REGION Network 17: Close Command
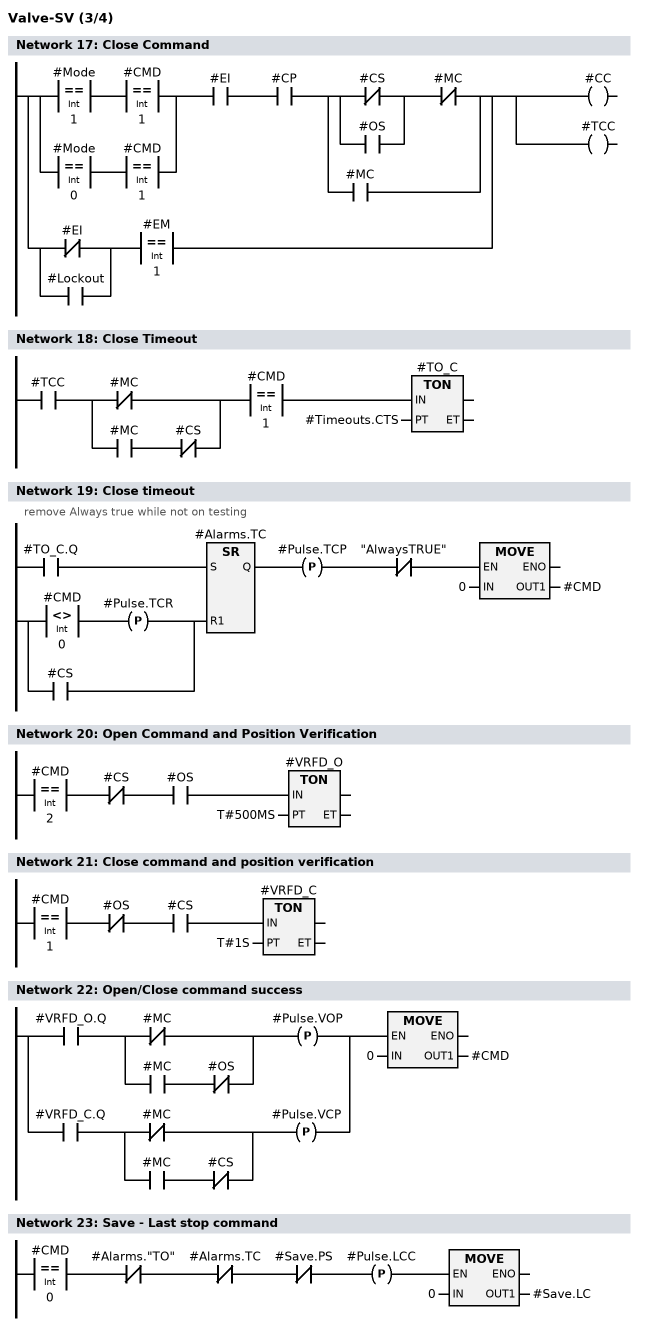
   RUNG wire#powerrail
      { S7_Templates := "SrcType := Int" } EQ_Contact(in1 := #Mode, in2 := 1)
      { S7_Templates := "SrcType := Int" } EQ_Contact(in1 := #CMD, in2 := 1)
      wire#w1
      Contact( #EI )
      Contact( #CP )
      wire#w2
      I_Contact( #CS )
      wire#w3
      I_Contact( #MC )
      wire#w4
      Coil( #CC )
   END_RUNG
   RUNG wire#powerrail
      { S7_Templates := "SrcType := Int" } EQ_Contact(in1 := #Mode, in2 := 0)
      { S7_Templates := "SrcType := Int" } EQ_Contact(in1 := #CMD, in2 := 1)
   END_RUNG wire#w1
   RUNG wire#w2
      Contact( #OS )
   END_RUNG wire#w3
   RUNG wire#w2
      Contact( #MC )
   END_RUNG wire#w4
   RUNG wire#powerrail
      I_Contact( #EI )
      wire#w5
      { S7_Templates := "SrcType := Int" } EQ_Contact(in1 := #EM, in2 := 1)
   END_RUNG wire#w4
   RUNG wire#powerrail
      Contact( #Lockout )
   END_RUNG wire#w5
   RUNG wire#w4
      Coil( #TCC )
   END_RUNG
   // the same network as SCL:
   #CC := ((((#Mode = 1) AND (#CMD = 1)) OR ((#Mode = 0) AND (#CMD = 1))) AND #EI AND #CP AND (((NOT #CS OR #OS) AND NOT #MC) OR #MC)) OR ((NOT #EI OR #Lockout) AND (#EM = 1));
   #TCC := #CC;
END_REGION

REGION Network 18: Close Timeout
   #TO_C(IN := #TCC AND (NOT #MC OR (#MC AND NOT #CS)) AND (#CMD = 1), PT := #Timeouts.CTS);   // TON
END_REGION

REGION Network 19: Close timeout
   // remove Always true while not on testing
   RUNG wire#powerrail
      Contact( #TO_C.Q )
      S_SR(operand := #Alarms.TC, r1 := wire#w1)
      P_Trig( #Pulse.TCP )
      I_Contact( "AlwaysTRUE" )
      { S7_GenerateENO := "TRUE" } Move(in := 0, out1 => #CMD)
   END_RUNG
   RUNG wire#powerrail
      { S7_Templates := "SrcType := Int" } NE_Contact(in1 := #CMD, in2 := 0)
      P_Trig( #Pulse.TCR )
   END_RUNG wire#w1
   RUNG wire#powerrail
      Contact( #CS )
   END_RUNG wire#w1
   // the same network as SCL:
   #_w1 := #CMD <> 0;
   #_w2 := #_w1 AND NOT #Pulse.TCR;   // rising edge
   #Pulse.TCR := #_w1;
   IF #TO_C.Q THEN
       #Alarms.TC := TRUE;   // SR flip-flop
   END_IF;
   IF #_w2 OR #CS THEN #Alarms.TC := FALSE; END_IF;
   #_w3 := #Alarms.TC AND NOT #Pulse.TCP;   // rising edge
   #Pulse.TCP := #Alarms.TC;
   IF #_w3 AND NOT "AlwaysTRUE" THEN #CMD := 0; END_IF;
END_REGION

REGION Network 20: Open Command and Position Verification
   #VRFD_O(IN := (#CMD = 2) AND NOT #CS AND #OS, PT := T#500MS);   // TON
END_REGION

REGION Network 21: Close command and position verification
   #VRFD_C(IN := (#CMD = 1) AND NOT #OS AND #CS, PT := T#1S);   // TON
END_REGION

REGION Network 22: Open/Close command success
   RUNG wire#powerrail
      Contact( #VRFD_O.Q )
      wire#w1
      I_Contact( #MC )
      wire#w2
      P_Trig( #Pulse.VOP )
      wire#w3
      { S7_GenerateENO := "TRUE" } Move(in := 0, out1 => #CMD)
   END_RUNG
   RUNG wire#w1
      Contact( #MC )
      I_Contact( #OS )
   END_RUNG wire#w2
   RUNG wire#powerrail
      Contact( #VRFD_C.Q )
      wire#w4
      I_Contact( #MC )
      wire#w5
      P_Trig( #Pulse.VCP )
   END_RUNG wire#w3
   RUNG wire#w4
      Contact( #MC )
      I_Contact( #CS )
   END_RUNG wire#w5
   // the same network as SCL:
   #_w1 := #VRFD_O.Q AND (NOT #MC OR (#MC AND NOT #OS));
   #_w2 := #_w1 AND NOT #Pulse.VOP;   // rising edge
   #Pulse.VOP := #_w1;
   #_w3 := #VRFD_C.Q AND (NOT #MC OR (#MC AND NOT #CS));
   #_w4 := #_w3 AND NOT #Pulse.VCP;   // rising edge
   #Pulse.VCP := #_w3;
   IF #_w2 OR #_w4 THEN #CMD := 0; END_IF;
END_REGION

REGION Network 23: Save - Last stop command
   RUNG wire#powerrail
      { S7_Templates := "SrcType := Int" } EQ_Contact(in1 := #CMD, in2 := 0)
      I_Contact( #Alarms."TO" )
      I_Contact( #Alarms.TC )
      I_Contact( #Save.PS )
      P_Trig( #Pulse.LCC )
      { S7_GenerateENO := "TRUE" } Move(in := 0, out1 => #Save.LC)
   END_RUNG
   // the same network as SCL:
   #_w1 := (#CMD = 0) AND NOT #Alarms."TO" AND NOT #Alarms.TC AND NOT #Save.PS;
   #_w2 := #_w1 AND NOT #Pulse.LCC;   // rising edge
   #Pulse.LCC := #_w1;
   IF #_w2 THEN #Save.LC := 0; END_IF;
END_REGION

REGION Network 24: Save - Last Stop Command
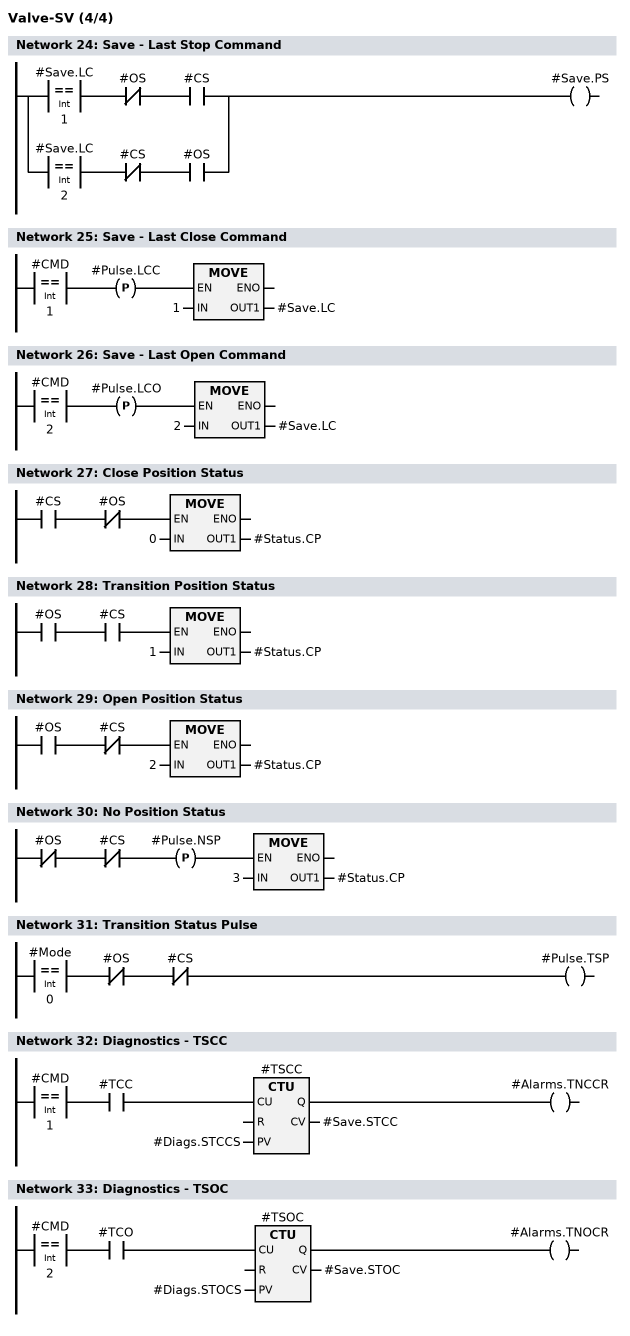
   RUNG wire#powerrail
      { S7_Templates := "SrcType := Int" } EQ_Contact(in1 := #Save.LC, in2 := 1)
      I_Contact( #OS )
      Contact( #CS )
      wire#w1
      Coil( #Save.PS )
   END_RUNG
   RUNG wire#powerrail
      { S7_Templates := "SrcType := Int" } EQ_Contact(in1 := #Save.LC, in2 := 2)
      I_Contact( #CS )
      Contact( #OS )
   END_RUNG wire#w1
   // the same network as SCL:
   #Save.PS := ((#Save.LC = 1) AND NOT #OS AND #CS) OR ((#Save.LC = 2) AND NOT #CS AND #OS);
END_REGION

REGION Network 25: Save - Last Close Command
   RUNG wire#powerrail
      { S7_Templates := "SrcType := Int" } EQ_Contact(in1 := #CMD, in2 := 1)
      P_Trig( #Pulse.LCC )
      { S7_GenerateENO := "TRUE" } Move(in := 1, out1 => #Save.LC)
   END_RUNG
   // the same network as SCL:
   #_w1 := #CMD = 1;
   #_w2 := #_w1 AND NOT #Pulse.LCC;   // rising edge
   #Pulse.LCC := #_w1;
   IF #_w2 THEN #Save.LC := 1; END_IF;
END_REGION

REGION Network 26: Save - Last Open Command
   RUNG wire#powerrail
      { S7_Templates := "SrcType := Int" } EQ_Contact(in1 := #CMD, in2 := 2)
      P_Trig( #Pulse.LCO )
      { S7_GenerateENO := "TRUE" } Move(in := 2, out1 => #Save.LC)
   END_RUNG
   // the same network as SCL:
   #_w1 := #CMD = 2;
   #_w2 := #_w1 AND NOT #Pulse.LCO;   // rising edge
   #Pulse.LCO := #_w1;
   IF #_w2 THEN #Save.LC := 2; END_IF;
END_REGION

REGION Network 27: Close Position Status
   RUNG wire#powerrail
      Contact( #CS )
      I_Contact( #OS )
      { S7_GenerateENO := "TRUE" } Move(in := 0, out1 => #Status.CP)
   END_RUNG
   // the same network as SCL:
   IF #CS AND NOT #OS THEN #Status.CP := 0; END_IF;
END_REGION

REGION Network 28: Transition Position Status
   RUNG wire#powerrail
      Contact( #OS )
      Contact( #CS )
      { S7_GenerateENO := "TRUE" } Move(in := 1, out1 => #Status.CP)
   END_RUNG
   // the same network as SCL:
   IF #OS AND #CS THEN #Status.CP := 1; END_IF;
END_REGION

REGION Network 29: Open Position Status
   RUNG wire#powerrail
      Contact( #OS )
      I_Contact( #CS )
      { S7_GenerateENO := "TRUE" } Move(in := 2, out1 => #Status.CP)
   END_RUNG
   // the same network as SCL:
   IF #OS AND NOT #CS THEN #Status.CP := 2; END_IF;
END_REGION

REGION Network 30: No Position Status
   RUNG wire#powerrail
      I_Contact( #OS )
      I_Contact( #CS )
      P_Trig( #Pulse.NSP )
      { S7_GenerateENO := "TRUE" } Move(in := 3, out1 => #Status.CP)
   END_RUNG
   // the same network as SCL:
   #_w1 := NOT #OS AND NOT #CS;
   #_w2 := #_w1 AND NOT #Pulse.NSP;   // rising edge
   #Pulse.NSP := #_w1;
   IF #_w2 THEN #Status.CP := 3; END_IF;
END_REGION

REGION Network 31: Transition Status Pulse
   RUNG wire#powerrail
      { S7_Templates := "SrcType := Int" } EQ_Contact(in1 := #Mode, in2 := 0)
      I_Contact( #OS )
      I_Contact( #CS )
      Coil( #Pulse.TSP )
   END_RUNG
   // the same network as SCL:
   #Pulse.TSP := (#Mode = 0) AND NOT #OS AND NOT #CS;
END_REGION

REGION Network 32: Diagnostics - TSCC
   #TSCC(CU := (#CMD = 1) AND #TCC, PV := #Diags.STCCS, CV => #Save.STCC);   // CTU
   #Alarms.TNCCR := #TSCC.Q;
END_REGION

REGION Network 33: Diagnostics - TSOC
   #TSOC(CU := (#CMD = 2) AND #TCO, PV := #Diags.STOCS, CV => #Save.STOC);   // CTU
   #Alarms.TNOCR := #TSOC.Q;
END_REGION
END_FUNCTION_BLOCK

FUNCTION_BLOCK "Valve-CV"   // FB801, LAD
TITLE = Valve-CV
{ S7_Optimized_Access := 'TRUE' }
VERSION : 0.1
// V1.0    GE    04/04/2022     Modified Unscale block and made sure CMD outputs right number.
   VAR_INPUT
      POS_CMD_Word : Word;   // Command in Word
      POS_FB : Int;   // Valve Position Raw Value
      AnalogFeedbackExists : Bool;   // Feedback Mode FALSE=FDBK Off // TRUE=FDBCK On
   END_VAR
   VAR_OUTPUT
      CMD : Int;   // Commanded Position in INT format
      CMD_R : Real;
   END_VAR
   VAR
      HMI : Struct
         Controls : Struct   // Controls
            SP : Real;   // Operator Command
            Lockout : Bool;
         END_STRUCT;
         Status : Struct   // Status
            POS : Real;   // Valve Position
            LST_POS : Real;   // Valve Position after a successful transition
            CMD_SP : Real;   // Commanded Position
            WR : Bool;   // Within Range
            UR_DB : Real;   // Upper range deadband
            LR_DB : Real;   // Lower range Deadband
            Mode_A : Bool;
            Mode_B : Bool;
         END_STRUCT;
         Alarms : Struct
            FCMD : Bool;   // SP vs PV mismatch timeout
            SP : Real;   // Setpoint Alarm (Unused)
            Error : Word;   // Unscaling Error
            IL : Bool := TRUE ;   // INTERLOCK (TRUE= GOOD FALSE = BAD)
         END_STRUCT;
         Config : Struct
            Mode : Int;   // 0 = PLC, 1 = HMI
            FDBK_MD : Int;   // Feedback Mode 0=FDBK Off // 1=FDBCK On
            WR_DB_TON : Time := T#1S;   // PV within range of SP
            WR_DB_TOF : Time := T#1S;   // PV within range of SP
            CMD_TO_TON_PT : Time := T#10S;   // Command to Open TON Preset Time
            CMD_TO_TOF_PT : Time := T#1S;   // Command to Open TOF Preset Time
            UR_DB_SP : Real := 1.0;   // Upper Range Deadband Setpoint
            LR_DB_SP : Real := 1.0;   // Lower Range Deadband Setpoint
            Min : Real;   // Minimum Output
            Max : Real := 100.0;   // Max Output
            failOpen : Bool;   // Enable Bipolar Values in Control Value
         END_STRUCT;
      END_STRUCT;
      OS : Struct
         SaveLastSP : Bool;   // Save Last Valid Setpoint
      END_STRUCT;
      WR_DB_TON : TON_TIME;   // Within Range Debounce TON
      WR_DB_TOF : TOF_TIME;   // Withing Range Debounce TOF
      CMD_TO_TON : TON_TIME;   // Command Timeout Debounce
      CMD_TO_TOF : TOF_TIME;   // Command Timeout Debounce
      "Lockout Trig" : Bool;
   END_VAR
   VAR_TEMP
      Scale : Struct
         RAI : Real;   // CV Position in REAL data type format
         EMax : Real;   // Engineering Max
         EMin : Real;   // Engineering Min
         RMax : Real;   // Raw Max
         RMin : Real;   // Raw Max
         OFST : Real;   // Offset
         RRAnge : Real;   // Raw Range
         ERange : Real;   // Engineering Range
      END_STRUCT;
      RDI : DInt;
      M1 : Real;
      M2 : Real;
      M3 : Real;
      CMD_SP : Real;
      WR : Bool;
      WR_DB : Bool;
      FCMD : Bool;   // SP vs PV mismatch timeout
      bypass : Bool;
      NRAIR : Real;
   END_VAR
   VAR_TEMP   // added for the SCL form of the ladder/FBD networks
      _w1 : Bool;
   END_VAR
BEGIN

REGION Network 1: Feedback MODE
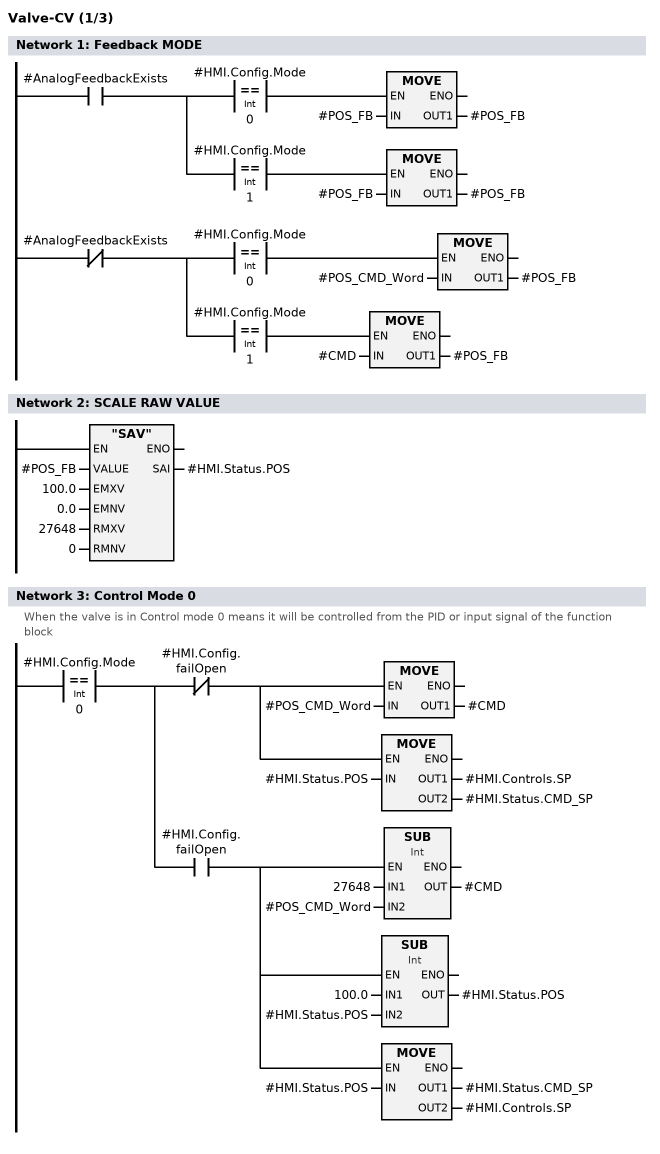
   RUNG wire#powerrail
      Contact( #AnalogFeedbackExists )
      wire#w1
      { S7_Templates := "SrcType := Int" } EQ_Contact(in1 := #HMI.Config.Mode, in2 := 0)
      Move(in := #POS_FB, out1 => #POS_FB)
   END_RUNG
   RUNG wire#w1
      { S7_Templates := "SrcType := Int" } EQ_Contact(in1 := #HMI.Config.Mode, in2 := 1)
      Move(in := #POS_FB, out1 => #POS_FB)
   END_RUNG
   RUNG wire#powerrail
      I_Contact( #AnalogFeedbackExists )
      wire#w2
      { S7_Templates := "SrcType := Int" } EQ_Contact(in1 := #HMI.Config.Mode, in2 := 0)
      Move(in := #POS_CMD_Word, out1 => #POS_FB)
   END_RUNG
   RUNG wire#w2
      { S7_Templates := "SrcType := Int" } EQ_Contact(in1 := #HMI.Config.Mode, in2 := 1)
      Move(in := #CMD, out1 => #POS_FB)
   END_RUNG
   // the same network as SCL:
   IF #AnalogFeedbackExists AND (#HMI.Config.Mode = 0) THEN #POS_FB := #POS_FB; END_IF;
   IF #AnalogFeedbackExists AND (#HMI.Config.Mode = 1) THEN #POS_FB := #POS_FB; END_IF;
   #_w1 := NOT #AnalogFeedbackExists;
   IF #_w1 AND (#HMI.Config.Mode = 0) THEN #POS_FB := #POS_CMD_Word; END_IF;
   IF #_w1 AND (#HMI.Config.Mode = 1) THEN #POS_FB := #CMD; END_IF;
END_REGION

REGION Network 2: SCALE RAW VALUE
   RUNG wire#powerrail
      "SAV"(VALUE := #POS_FB, EMXV := 100.0, EMNV := 0.0, RMXV := 27648, RMNV := 0, SAI => #HMI.Status.POS)
   END_RUNG
   // the same network as SCL:
   "SAV"(VALUE := #POS_FB, EMXV := 100.0, EMNV := 0.0, RMXV := 27648, RMNV := 0, SAI => #HMI.Status.POS);
END_REGION

REGION Network 3: Control Mode 0
   // When the valve is in Control mode 0 means it will be controlled from the PID or input signal of the function block
   RUNG wire#powerrail
      { S7_Templates := "SrcType := Int" } EQ_Contact(in1 := #HMI.Config.Mode, in2 := 0)
      wire#w1
      I_Contact( #HMI.Config.failOpen )
      wire#w2
      { S7_GenerateENO := "TRUE" } Move(in := #POS_CMD_Word, out1 => #CMD)
   END_RUNG
   RUNG wire#w2
      Move(in := #HMI.Status.POS, out1 => #HMI.Controls.SP, out2 => #HMI.Status.CMD_SP)
   END_RUNG
   RUNG wire#w1
      Contact( #HMI.Config.failOpen )
      wire#w3
      { S7_Templates := "SrcType := Int" } Sub(in1 := 27648, in2 := #POS_CMD_Word, out => #CMD)
   END_RUNG
   RUNG wire#w3
      { S7_Templates := "SrcType := Int" } Sub(in1 := 100.0, in2 := #HMI.Status.POS, out => #HMI.Status.POS)
   END_RUNG
   RUNG wire#w3
      Move(in := #HMI.Status.POS, out1 => #HMI.Status.CMD_SP, out2 => #HMI.Controls.SP)
   END_RUNG
   // the same network as SCL:
   #_w1 := #HMI.Config.Mode = 0;
   IF #_w1 AND NOT #HMI.Config.failOpen THEN
       #CMD := #POS_CMD_Word;
       #HMI.Controls.SP := #HMI.Status.POS;
       #HMI.Status.CMD_SP := #HMI.Status.POS;
   END_IF;
   IF #_w1 AND #HMI.Config.failOpen THEN
       #CMD := 27648 - #POS_CMD_Word;
       #HMI.Status.POS := 100.0 - #HMI.Status.POS;
       #HMI.Status.CMD_SP := #HMI.Status.POS;
       #HMI.Controls.SP := #HMI.Status.POS;
   END_IF;
END_REGION

REGION Network 4: Control Mode 1
   // Control Mode 1 will control from HMI (force valve to go to a certain position)
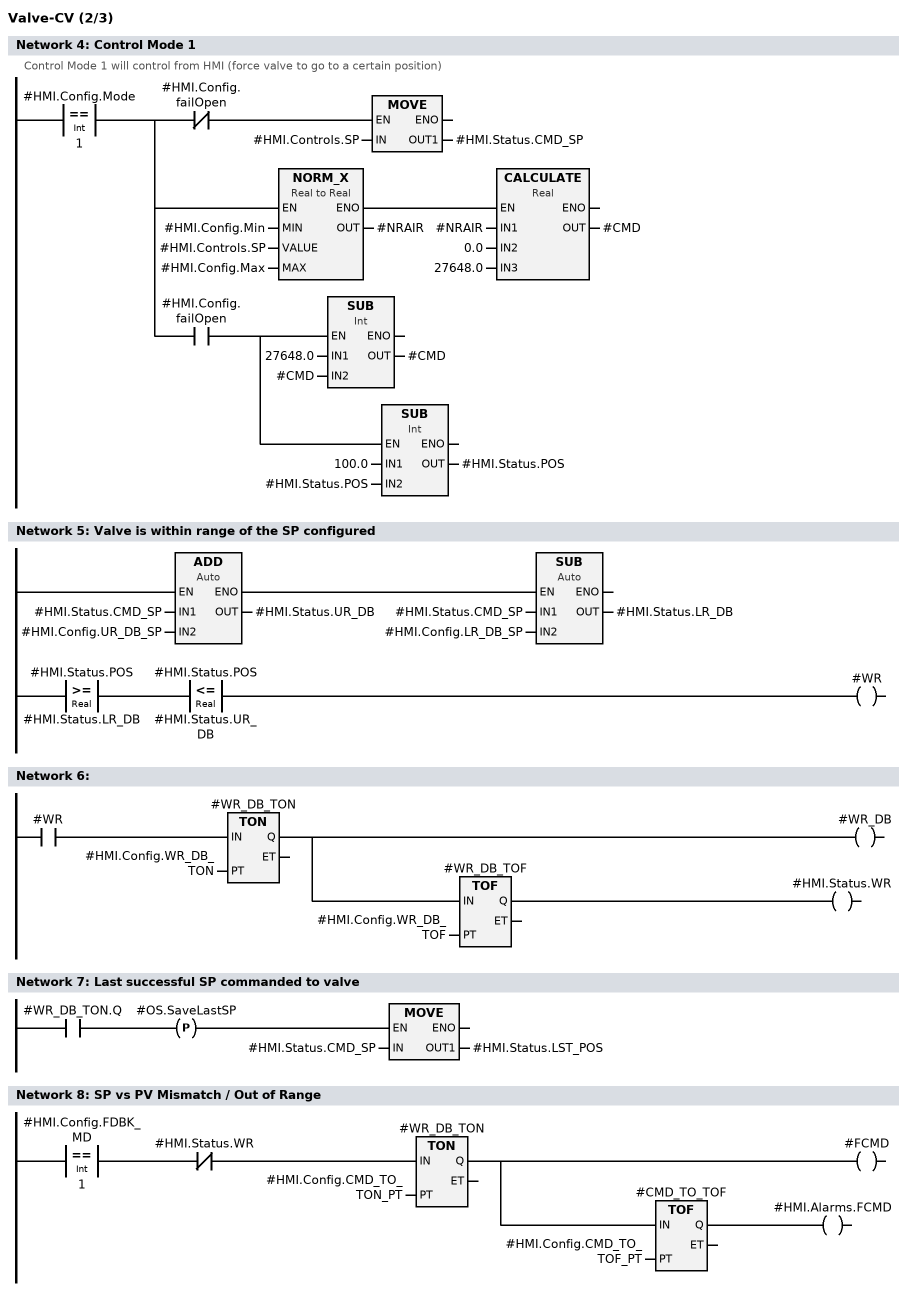
   RUNG wire#powerrail
      { S7_Templates := "SrcType := Int" } EQ_Contact(in1 := #HMI.Config.Mode, in2 := 1)
      wire#w1
      I_Contact( #HMI.Config.failOpen )
      { S7_GenerateENO := "TRUE" } Move(in := #HMI.Controls.SP, out1 => #HMI.Status.CMD_SP)
   END_RUNG
   RUNG wire#w1
      { S7_Templates := "[SrcType := Real, DestType := Real]" } Normalize(min := #HMI.Config.Min, value := #HMI.Controls.SP, max := #HMI.Config.Max, out => #NRAIR)
      { S7_Templates := "SrcType := Real"; S7_Expression := "(IN1 * (IN3 - IN2)) + IN2" } Calculate(in1 := #NRAIR, in2 := 0.0, in3 := 27648.0, out => #CMD)
   END_RUNG
   RUNG wire#w1
      Contact( #HMI.Config.failOpen )
      wire#w2
      { S7_Templates := "SrcType := Int" } Sub(in1 := 27648.0, in2 := #CMD, out => #CMD)
   END_RUNG
   RUNG wire#w2
      { S7_Templates := "SrcType := Int" } Sub(in1 := 100.0, in2 := #HMI.Status.POS, out => #HMI.Status.POS)
   END_RUNG
   // the same network as SCL:
   #_w1 := #HMI.Config.Mode = 1;
   IF #_w1 AND NOT #HMI.Config.failOpen THEN #HMI.Status.CMD_SP := #HMI.Controls.SP; END_IF;
   IF #_w1 THEN
       #NRAIR := NORM_X(MIN := #HMI.Config.Min, VALUE := #HMI.Controls.SP, MAX := #HMI.Config.Max);
       #CMD := (#NRAIR * (27648.0 - 0.0)) + 0.0;
   END_IF;
   IF #_w1 AND #HMI.Config.failOpen THEN
       #CMD := 27648.0 - #CMD;
       #HMI.Status.POS := 100.0 - #HMI.Status.POS;
   END_IF;
END_REGION

REGION Network 5: Valve is within range of the SP configured
   RUNG wire#powerrail
      Add(in1 := #HMI.Status.CMD_SP, in2 := #HMI.Config.UR_DB_SP, out => #HMI.Status.UR_DB)
      Sub(in1 := #HMI.Status.CMD_SP, in2 := #HMI.Config.LR_DB_SP, out => #HMI.Status.LR_DB)
   END_RUNG
   RUNG wire#powerrail
      { S7_Templates := "SrcType := Real" } GE_Contact(in1 := #HMI.Status.POS, in2 := #HMI.Status.LR_DB)
      { S7_Templates := "SrcType := Real" } LE_Contact(in1 := #HMI.Status.POS, in2 := #HMI.Status.UR_DB)
      Coil( #WR )
   END_RUNG
   // the same network as SCL:
   #HMI.Status.UR_DB := #HMI.Status.CMD_SP + #HMI.Config.UR_DB_SP;
   #HMI.Status.LR_DB := #HMI.Status.CMD_SP - #HMI.Config.LR_DB_SP;
   #WR := (#HMI.Status.POS >= #HMI.Status.LR_DB) AND (#HMI.Status.POS <= #HMI.Status.UR_DB);
END_REGION

REGION Network 6
   #WR_DB_TON(IN := #WR, PT := #HMI.Config.WR_DB_TON);   // TON
   #WR_DB := #WR_DB_TON.Q;
   #WR_DB_TOF(IN := #WR_DB_TON.Q, PT := #HMI.Config.WR_DB_TOF);   // TOF
   #HMI.Status.WR := #WR_DB_TOF.Q;
END_REGION

REGION Network 7: Last successful SP commanded to valve
   RUNG wire#powerrail
      Contact( #WR_DB_TON.Q )
      P_Trig( #OS.SaveLastSP )
      { S7_GenerateENO := "TRUE" } Move(in := #HMI.Status.CMD_SP, out1 => #HMI.Status.LST_POS)
   END_RUNG
   // the same network as SCL:
   #_w1 := #WR_DB_TON.Q AND NOT #OS.SaveLastSP;   // rising edge
   #OS.SaveLastSP := #WR_DB_TON.Q;
   IF #_w1 THEN #HMI.Status.LST_POS := #HMI.Status.CMD_SP; END_IF;
END_REGION

REGION Network 8: SP vs PV Mismatch / Out of Range
   #WR_DB_TON(IN := (#HMI.Config.FDBK_MD = 1) AND NOT #HMI.Status.WR, PT := #HMI.Config.CMD_TO_TON_PT);   // TON
   #FCMD := #WR_DB_TON.Q;
   #CMD_TO_TOF(IN := #WR_DB_TON.Q, PT := #HMI.Config.CMD_TO_TOF_PT);   // TOF
   #HMI.Alarms.FCMD := #CMD_TO_TOF.Q;
END_REGION

REGION Network 9: Lockout Sequence
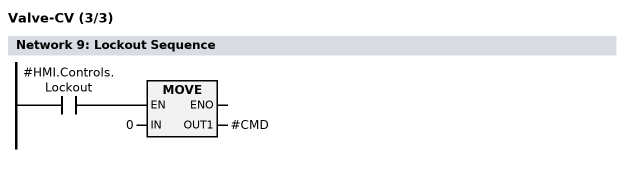
   RUNG wire#powerrail
      Contact( #HMI.Controls.Lockout )
      { S7_GenerateENO := "TRUE" } Move(in := 0, out1 => #CMD)
   END_RUNG
   // the same network as SCL:
   IF #HMI.Controls.Lockout THEN #CMD := 0; END_IF;
END_REGION
END_FUNCTION_BLOCK

// folder: Analogs inputs

FUNCTION "Analog Trasmitter" : Void   // FC5, LAD
TITLE = Analog Trasmitter Fuction Code
{ S7_Optimized_Access := 'TRUE' }
VERSION : 0.1
// Updated Date:
// Note:
BEGIN
END_FUNCTION

// folder: Analogs inputs/Trasmitters/Analyzer Trasmitters

FUNCTION "Analyzer Trasmitters" : Void   // FC16, LAD
TITLE = Analyzer Trasmitters
{ S7_Optimized_Access := 'TRUE' }
VERSION : 0.1
// Updated Date:
// Note:
BEGIN

REGION Network 1: AT-3011 : C-301 Nitrates Analyzer #1
   // Erick
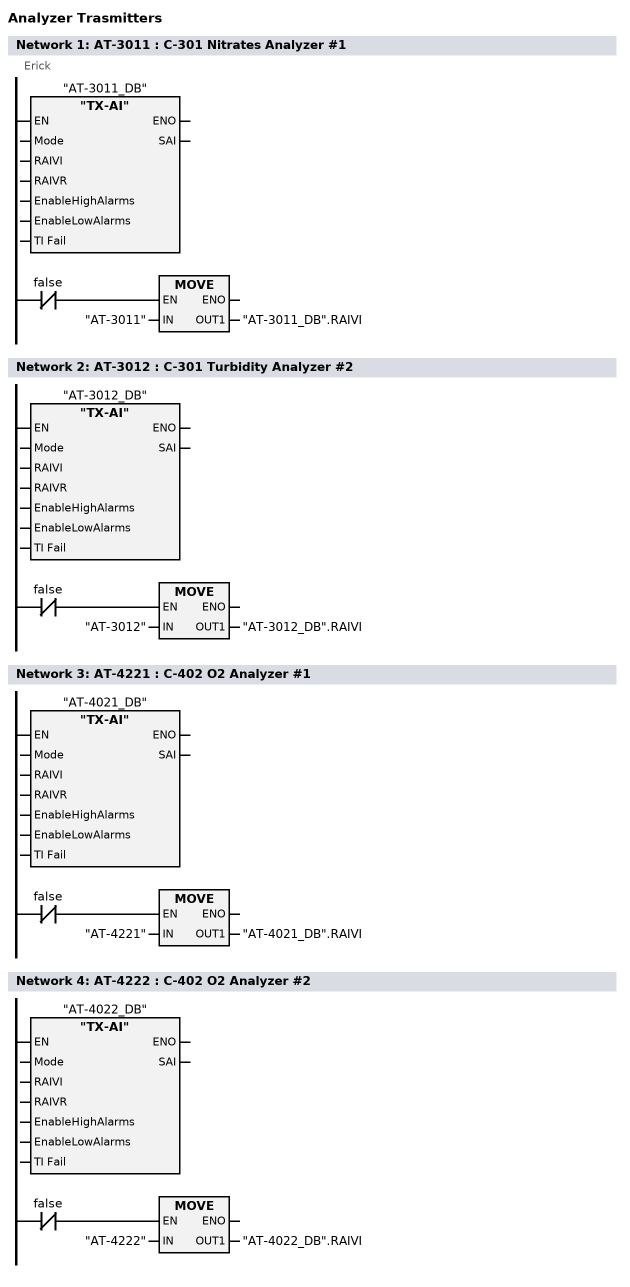
   RUNG wire#powerrail
      "AT-3011_DB"(Mode :=, RAIVI :=, RAIVR :=, EnableHighAlarms :=, EnableLowAlarms :=, "TI Fail" :=, SAI =>)
   END_RUNG
   RUNG wire#powerrail
      I_Contact( false )
      { S7_GenerateENO := "TRUE" } Move(in := "AT-3011", out1 => "AT-3011_DB".RAIVI)
   END_RUNG
   // the same network as SCL:
   "AT-3011_DB"();   // "TX-AI"
   IF NOT false THEN "AT-3011_DB".RAIVI := "AT-3011"; END_IF;
END_REGION

REGION Network 2: AT-3012 : C-301 Turbidity Analyzer #2
   RUNG wire#powerrail
      "AT-3012_DB"(Mode :=, RAIVI :=, RAIVR :=, EnableHighAlarms :=, EnableLowAlarms :=, "TI Fail" :=, SAI =>)
   END_RUNG
   RUNG wire#powerrail
      I_Contact( false )
      { S7_GenerateENO := "TRUE" } Move(in := "AT-3012", out1 => "AT-3012_DB".RAIVI)
   END_RUNG
   // the same network as SCL:
   "AT-3012_DB"();   // "TX-AI"
   IF NOT false THEN "AT-3012_DB".RAIVI := "AT-3012"; END_IF;
END_REGION

REGION Network 3: AT-4221 : C-402 O2 Analyzer #1
   RUNG wire#powerrail
      "AT-4021_DB"(Mode :=, RAIVI :=, RAIVR :=, EnableHighAlarms :=, EnableLowAlarms :=, "TI Fail" :=, SAI =>)
   END_RUNG
   RUNG wire#powerrail
      I_Contact( false )
      { S7_GenerateENO := "TRUE" } Move(in := "AT-4221", out1 => "AT-4021_DB".RAIVI)
   END_RUNG
   // the same network as SCL:
   "AT-4021_DB"();   // "TX-AI"
   IF NOT false THEN "AT-4021_DB".RAIVI := "AT-4221"; END_IF;
END_REGION

REGION Network 4: AT-4222 : C-402 O2 Analyzer #2
   RUNG wire#powerrail
      "AT-4022_DB"(Mode :=, RAIVI :=, RAIVR :=, EnableHighAlarms :=, EnableLowAlarms :=, "TI Fail" :=, SAI =>)
   END_RUNG
   RUNG wire#powerrail
      I_Contact( false )
      { S7_GenerateENO := "TRUE" } Move(in := "AT-4222", out1 => "AT-4022_DB".RAIVI)
   END_RUNG
   // the same network as SCL:
   "AT-4022_DB"();   // "TX-AI"
   IF NOT false THEN "AT-4022_DB".RAIVI := "AT-4222"; END_IF;
END_REGION
END_FUNCTION

// folder: Analogs inputs/Trasmitters/Flow Trasmitters

FUNCTION "FlowTrasmitters" : Void   // FC8, LAD
TITLE = Flow Trasmitter Fuction Code
{ S7_Optimized_Access := 'TRUE' }
VERSION : 0.1
// Updated Date:
// Note:
BEGIN

REGION Network 1: FT-1011: T-101 Recirc Flow
   // "FT-1011"
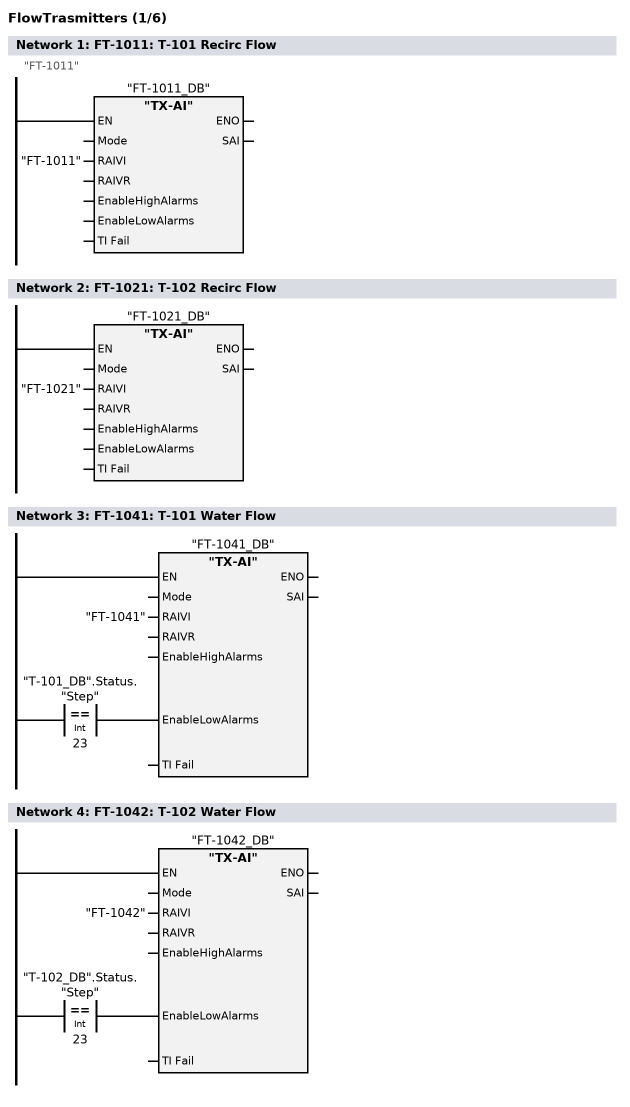
   RUNG wire#powerrail
      "FT-1011_DB"(Mode :=, RAIVI := "FT-1011", RAIVR :=, EnableHighAlarms :=, EnableLowAlarms :=, "TI Fail" :=, SAI =>)
   END_RUNG
   // the same network as SCL:
   "FT-1011_DB"(RAIVI := "FT-1011");   // "TX-AI"
END_REGION

REGION Network 2: FT-1021: T-102 Recirc Flow
   RUNG wire#powerrail
      "FT-1021_DB"(Mode :=, RAIVI := "FT-1021", RAIVR :=, EnableHighAlarms :=, EnableLowAlarms :=, "TI Fail" :=, SAI =>)
   END_RUNG
   // the same network as SCL:
   "FT-1021_DB"(RAIVI := "FT-1021");   // "TX-AI"
END_REGION

REGION Network 3: FT-1041: T-101 Water Flow
   RUNG wire#powerrail
      "FT-1041_DB"(EnableLowAlarms := wire#w1, Mode :=, RAIVI := "FT-1041", RAIVR :=, EnableHighAlarms :=, "TI Fail" :=, SAI =>)
   END_RUNG
   RUNG wire#powerrail
      { S7_Templates := "SrcType := Int" } EQ_Contact(in1 := "T-101_DB".Status."Step", in2 := 23)
   END_RUNG wire#w1
   // the same network as SCL:
   "FT-1041_DB"(RAIVI := "FT-1041", EnableLowAlarms := "T-101_DB".Status."Step" = 23);   // "TX-AI"
END_REGION

REGION Network 4: FT-1042: T-102 Water Flow
   RUNG wire#powerrail
      "FT-1042_DB"(EnableLowAlarms := wire#w1, Mode :=, RAIVI := "FT-1042", RAIVR :=, EnableHighAlarms :=, "TI Fail" :=, SAI =>)
   END_RUNG
   RUNG wire#powerrail
      { S7_Templates := "SrcType := Int" } EQ_Contact(in1 := "T-102_DB".Status."Step", in2 := 23)
   END_RUNG wire#w1
   // the same network as SCL:
   "FT-1042_DB"(RAIVI := "FT-1042", EnableLowAlarms := "T-102_DB".Status."Step" = 23);   // "TX-AI"
END_REGION

REGION Network 5: FT-1043:R-201 Water Flow
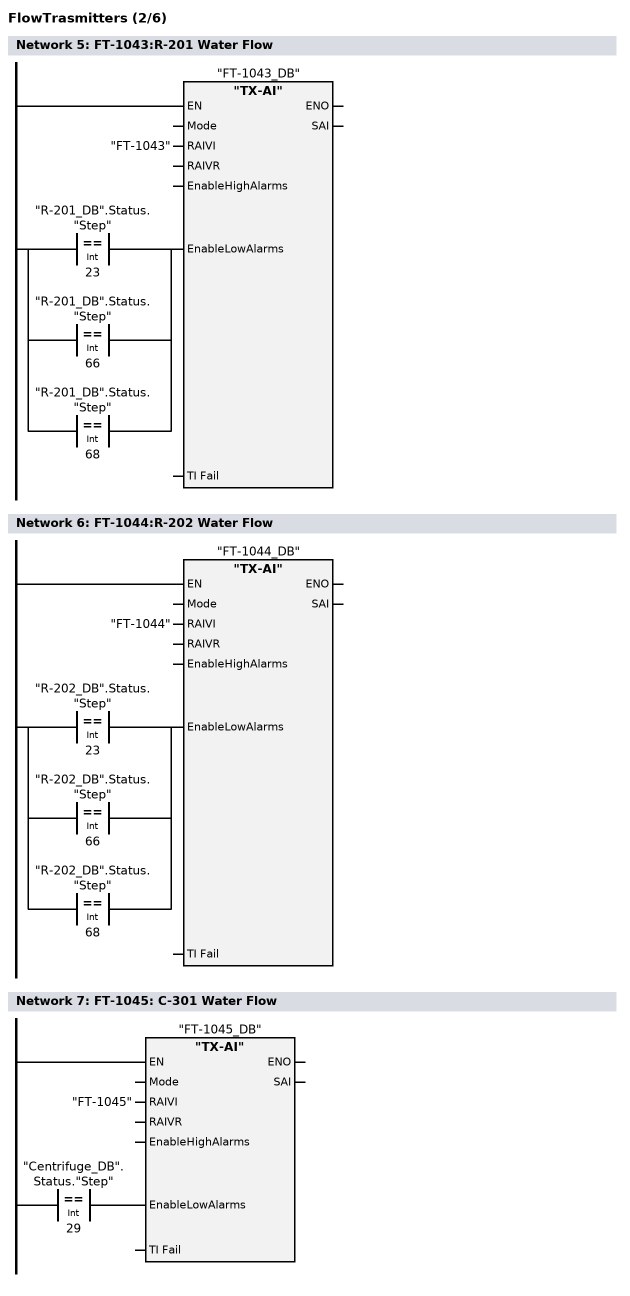
   RUNG wire#powerrail
      "FT-1043_DB"(EnableLowAlarms := wire#w1, Mode :=, RAIVI := "FT-1043", RAIVR :=, EnableHighAlarms :=, "TI Fail" :=, SAI =>)
   END_RUNG
   RUNG wire#powerrail
      { S7_Templates := "SrcType := Int" } EQ_Contact(in1 := "R-201_DB".Status."Step", in2 := 23)
   END_RUNG wire#w1
   RUNG wire#powerrail
      { S7_Templates := "SrcType := Int" } EQ_Contact(in1 := "R-201_DB".Status."Step", in2 := 66)
   END_RUNG wire#w1
   RUNG wire#powerrail
      { S7_Templates := "SrcType := Int" } EQ_Contact(in1 := "R-201_DB".Status."Step", in2 := 68)
   END_RUNG wire#w1
   // the same network as SCL:
   "FT-1043_DB"(RAIVI := "FT-1043",   // "TX-AI"
                EnableLowAlarms := ("R-201_DB".Status."Step" = 23) OR ("R-201_DB".Status."Step" = 66) OR ("R-201_DB".Status."Step" = 68));
END_REGION

REGION Network 6: FT-1044:R-202 Water Flow
   RUNG wire#powerrail
      "FT-1044_DB"(EnableLowAlarms := wire#w1, Mode :=, RAIVI := "FT-1044", RAIVR :=, EnableHighAlarms :=, "TI Fail" :=, SAI =>)
   END_RUNG
   RUNG wire#powerrail
      { S7_Templates := "SrcType := Int" } EQ_Contact(in1 := "R-202_DB".Status."Step", in2 := 23)
   END_RUNG wire#w1
   RUNG wire#powerrail
      { S7_Templates := "SrcType := Int" } EQ_Contact(in1 := "R-202_DB".Status."Step", in2 := 66)
   END_RUNG wire#w1
   RUNG wire#powerrail
      { S7_Templates := "SrcType := Int" } EQ_Contact(in1 := "R-202_DB".Status."Step", in2 := 68)
   END_RUNG wire#w1
   // the same network as SCL:
   "FT-1044_DB"(RAIVI := "FT-1044",   // "TX-AI"
                EnableLowAlarms := ("R-202_DB".Status."Step" = 23) OR ("R-202_DB".Status."Step" = 66) OR ("R-202_DB".Status."Step" = 68));
END_REGION

REGION Network 7: FT-1045: C-301 Water Flow
   RUNG wire#powerrail
      "FT-1045_DB"(EnableLowAlarms := wire#w1, Mode :=, RAIVI := "FT-1045", RAIVR :=, EnableHighAlarms :=, "TI Fail" :=, SAI =>)
   END_RUNG
   RUNG wire#powerrail
      { S7_Templates := "SrcType := Int" } EQ_Contact(in1 := "Centrifuge_DB".Status."Step", in2 := 29)
   END_RUNG wire#w1
   // the same network as SCL:
   "FT-1045_DB"(RAIVI := "FT-1045", EnableLowAlarms := "Centrifuge_DB".Status."Step" = 29);   // "TX-AI"
END_REGION

REGION Network 8: FT-2011:T-101 to R-201 Flow
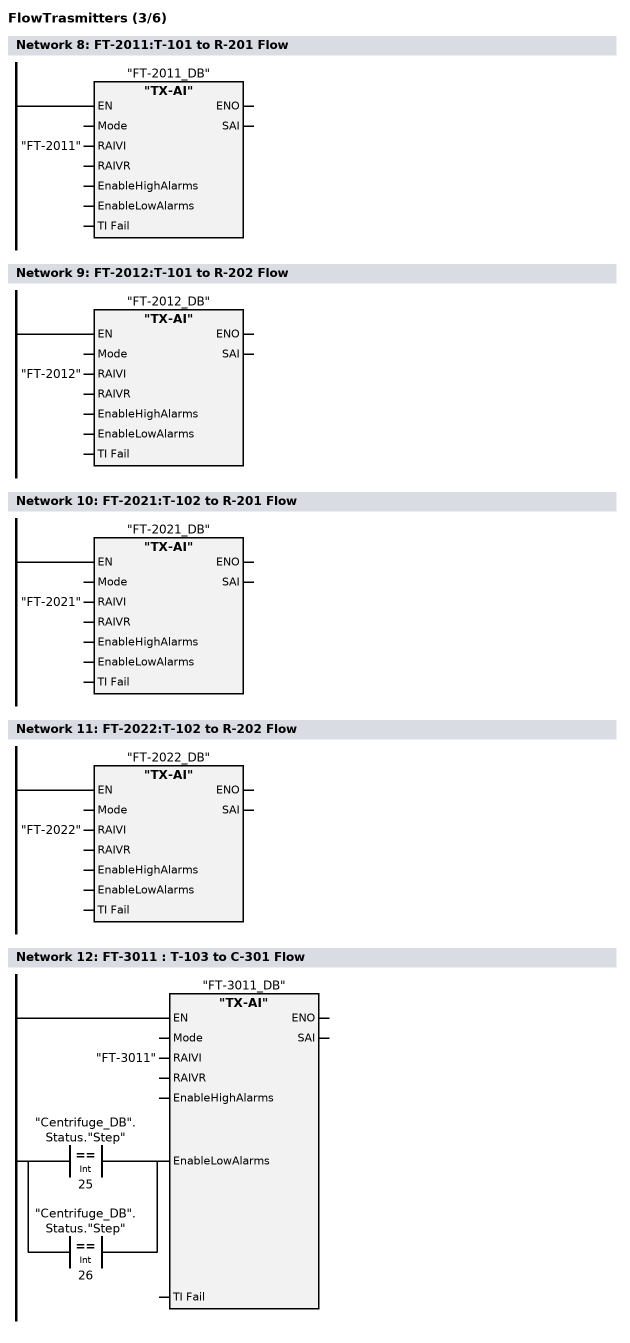
   RUNG wire#powerrail
      "FT-2011_DB"(Mode :=, RAIVI := "FT-2011", RAIVR :=, EnableHighAlarms :=, EnableLowAlarms :=, "TI Fail" :=, SAI =>)
   END_RUNG
   // the same network as SCL:
   "FT-2011_DB"(RAIVI := "FT-2011");   // "TX-AI"
END_REGION

REGION Network 9: FT-2012:T-101 to R-202 Flow
   RUNG wire#powerrail
      "FT-2012_DB"(Mode :=, RAIVI := "FT-2012", RAIVR :=, EnableHighAlarms :=, EnableLowAlarms :=, "TI Fail" :=, SAI =>)
   END_RUNG
   // the same network as SCL:
   "FT-2012_DB"(RAIVI := "FT-2012");   // "TX-AI"
END_REGION

REGION Network 10: FT-2021:T-102 to R-201 Flow
   RUNG wire#powerrail
      "FT-2021_DB"(Mode :=, RAIVI := "FT-2021", RAIVR :=, EnableHighAlarms :=, EnableLowAlarms :=, "TI Fail" :=, SAI =>)
   END_RUNG
   // the same network as SCL:
   "FT-2021_DB"(RAIVI := "FT-2021");   // "TX-AI"
END_REGION

REGION Network 11: FT-2022:T-102 to R-202 Flow
   RUNG wire#powerrail
      "FT-2022_DB"(Mode :=, RAIVI := "FT-2022", RAIVR :=, EnableHighAlarms :=, EnableLowAlarms :=, "TI Fail" :=, SAI =>)
   END_RUNG
   // the same network as SCL:
   "FT-2022_DB"(RAIVI := "FT-2022");   // "TX-AI"
END_REGION

REGION Network 12: FT-3011 : T-103 to C-301 Flow
   RUNG wire#powerrail
      "FT-3011_DB"(EnableLowAlarms := wire#w1, Mode :=, RAIVI := "FT-3011", RAIVR :=, EnableHighAlarms :=, "TI Fail" :=, SAI =>)
   END_RUNG
   RUNG wire#powerrail
      { S7_Templates := "SrcType := Int" } EQ_Contact(in1 := "Centrifuge_DB".Status."Step", in2 := 25)
   END_RUNG wire#w1
   RUNG wire#powerrail
      { S7_Templates := "SrcType := Int" } EQ_Contact(in1 := "Centrifuge_DB".Status."Step", in2 := 26)
   END_RUNG wire#w1
   // the same network as SCL:
   "FT-3011_DB"(RAIVI := "FT-3011",   // "TX-AI"
                EnableLowAlarms := ("Centrifuge_DB".Status."Step" = 25) OR ("Centrifuge_DB".Status."Step" = 26));
END_REGION

REGION Network 13: FT-3012: C-301 Outlet Flow
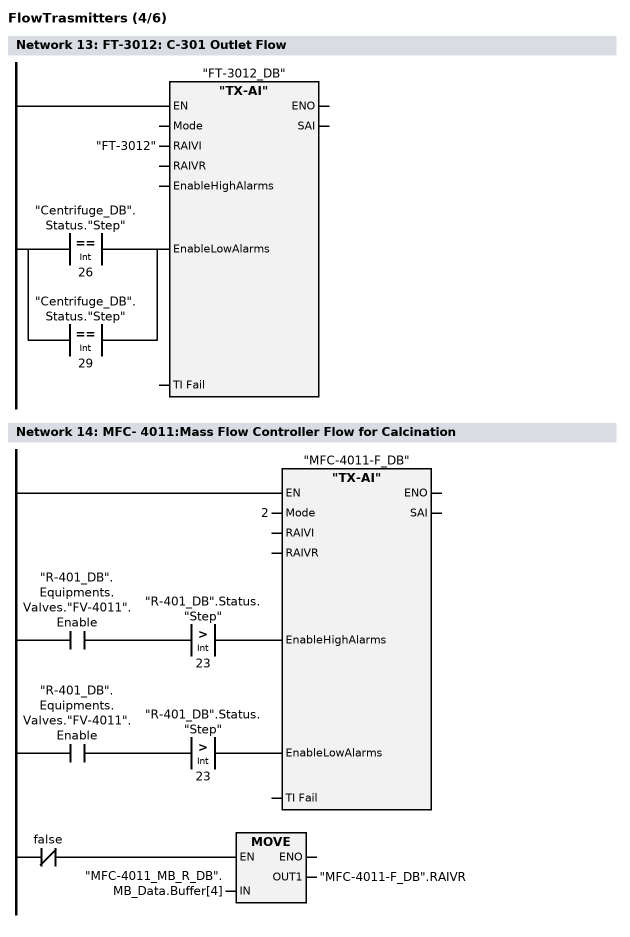
   RUNG wire#powerrail
      "FT-3012_DB"(EnableLowAlarms := wire#w1, Mode :=, RAIVI := "FT-3012", RAIVR :=, EnableHighAlarms :=, "TI Fail" :=, SAI =>)
   END_RUNG
   RUNG wire#powerrail
      { S7_Templates := "SrcType := Int" } EQ_Contact(in1 := "Centrifuge_DB".Status."Step", in2 := 26)
   END_RUNG wire#w1
   RUNG wire#powerrail
      { S7_Templates := "SrcType := Int" } EQ_Contact(in1 := "Centrifuge_DB".Status."Step", in2 := 29)
   END_RUNG wire#w1
   // the same network as SCL:
   "FT-3012_DB"(RAIVI := "FT-3012",   // "TX-AI"
                EnableLowAlarms := ("Centrifuge_DB".Status."Step" = 26) OR ("Centrifuge_DB".Status."Step" = 29));
END_REGION
